VERSION : 0.1
   VAR
      ReadWriteDeviceNo : Int := 0;
      CopyDeviceNO : Int := 0;
      Read : Bool := FALSE;
      Write : Bool := FALSE;
      Copy : Bool := FALSE;
      Tank : Array[0..12] of "UDT502_PV_Tank";
   END_VAR
BEGIN
   Tank[1].Level.PV_Conf_ActV.Address := 324;
   Tank[2].Level.PV_Conf_ActV.Address := 326;
   Tank[1].Level.PV_Conf_ActV.Multiplier := 10.0;
   Tank[2].Level.PV_Conf_ActV.Multiplier := 10.0;
   Tank[1].Level.PV_Conf_ActV.MaxValueSensor := 0.0;
   Tank[2].Level.PV_Conf_ActV.MaxValueSensor := 0.0;
   Tank[2].Level.PV_Conf_ActV.MinValueSensor := 0.0;
   Tank[1].Temp.PV_Conf_ActV.Address := 300;
   Tank[1].Level.PV_Conf_ActV.MinValueSensor := 0.0;
   Tank[2].Temp.PV_Conf_ActV.Address := 302;
   Tank[1].Temp.PV_Conf_ActV.Multiplier := 100.0;
   Tank[2].Temp.PV_Conf_ActV.Multiplier := 100.0;
   Tank[0].Temp.PV_SetV.Value := 15.0;
   Tank[0].Temp.PV_SetV.WarningLowerLimit := 0.0;
   Tank[0].Temp.PV_SetV.WarningUpperLimit := 0.0;
   Tank[0].Temp.PV_SetV.AlarmLowerLimit := 0.0;
   Tank[0].Temp.PV_SetV.AlarmUpperLimit := 0.0;
   Tank[0].Temp.PV_Conf_ActV.ModulNo := 1;
   Tank[0].Temp.PV_Conf_ActV.Address := 300;
   Tank[0].Temp.PV_Conf_ActV.OffsetSignal := 0;
   Tank[0].Temp.PV_Conf_ActV.Multiplier := 100.0;
   Tank[0].Temp.PV_Conf_ActV.MinValueSensor := 1.0;
   Tank[0].Temp.PV_Conf_ActV.MaxValueSensor := 10000.0;
   Tank[0].Temp.PV_Conf_ActV.MaxSignalResolution := 0.0;
   Tank[0].Level.PV_SetV.Value := 0.0;
   Tank[0].Level.PV_SetV.WarningLowerLimit := 0.0;
   Tank[0].Level.PV_SetV.WarningUpperLimit := 0.0;
   Tank[0].Level.PV_SetV.AlarmLowerLimit := 0.0;
   Tank[0].Level.PV_SetV.AlarmUpperLimit := 0.0;
   Tank[0].Level.PV_Conf_ActV.ModulNo := 1;
   Tank[0].Level.PV_Conf_ActV.Address := 324;
   Tank[0].Level.PV_Conf_ActV.OffsetSignal := 0;
   Tank[0].Level.PV_Conf_ActV.Multiplier := 10.0;
   Tank[0].Level.PV_Conf_ActV.MinValueSensor := 0.0;
   Tank[0].Level.PV_Conf_ActV.MaxValueSensor := 0.0;
   Tank[0].Level.PV_Conf_ActV.MaxSignalResolution := 0.0;
   Tank[0].Pressure.PV_SetV.Value := 0.0;
   Tank[0].Pressure.PV_SetV.WarningLowerLimit := 0.0;
   Tank[0].Pressure.PV_SetV.WarningUpperLimit := 0.0;
   Tank[0].Pressure.PV_SetV.AlarmLowerLimit := 0.0;
   Tank[0].Pressure.PV_SetV.AlarmUpperLimit := 0.0;
   Tank[0].Pressure.PV_Conf_ActV.ModulNo := 0;
   Tank[0].Pressure.PV_Conf_ActV.Address := 0;
   Tank[0].Pressure.PV_Conf_ActV.OffsetSignal := 0;
   Tank[0].Pressure.PV_Conf_ActV.Multiplier := 0.0;
   Tank[0].Pressure.PV_Conf_ActV.MinValueSensor := 0.0;
   Tank[0].Pressure.PV_Conf_ActV.MaxValueSensor := 0.0;
   Tank[0].Pressure.PV_Conf_ActV.MaxSignalResolution := 0.0;
   Tank[0].Nucleation.PV_SetV.Value := 2.0;
   Tank[0].Nucleation.PV_SetV.WarningLowerLimit := 0.0;
   Tank[0].Nucleation.PV_SetV.WarningUpperLimit := 0.0;
   Tank[0].Nucleation.PV_SetV.AlarmLowerLimit := 0.0;
   Tank[0].Nucleation.PV_SetV.AlarmUpperLimit := 0.0;
   Tank[0].Nucleation.PV_Conf_ActV.ModulNo := 1;
   Tank[0].Nucleation.PV_Conf_ActV.Address := 330;
   Tank[0].Nucleation.PV_Conf_ActV.OffsetSignal := 0;
   Tank[0].Nucleation.PV_Conf_ActV.Multiplier := 10.0;
   Tank[0].Nucleation.PV_Conf_ActV.MinValueSensor := 0.0;
   Tank[0].Nucleation.PV_Conf_ActV.MaxValueSensor := 100.0;
   Tank[0].Nucleation.PV_Conf_ActV.MaxSignalResolution := 0.0;
   Tank[0].JacketHeater.PV_SetV.Value := 0.0;
   Tank[0].JacketHeater.PV_SetV.WarningLowerLimit := 0.0;
   Tank[0].JacketHeater.PV_SetV.WarningUpperLimit := 0.0;
   Tank[0].JacketHeater.PV_SetV.AlarmLowerLimit := 0.0;
   Tank[0].JacketHeater.PV_SetV.AlarmUpperLimit := 0.0;
   Tank[0].JacketHeater.PV_Conf_ActV.ModulNo := 0;
   Tank[0].JacketHeater.PV_Conf_ActV.Address := 0;
   Tank[0].JacketHeater.PV_Conf_ActV.OffsetSignal := 0;
   Tank[0].JacketHeater.PV_Conf_ActV.Multiplier := 0.0;
   Tank[0].JacketHeater.PV_Conf_ActV.MinValueSensor := 0.0;
   Tank[0].JacketHeater.PV_Conf_ActV.MaxValueSensor := 0.0;
   Tank[0].JacketHeater.PV_Conf_ActV.MaxSignalResolution := 0.0;
   Tank[1].Temp.PV_SetV.Value := 15.0;
   Tank[1].Temp.PV_SetV.WarningLowerLimit := 0.0;
   Tank[1].Temp.PV_SetV.WarningUpperLimit := 0.0;
   Tank[1].Temp.PV_SetV.AlarmLowerLimit := 0.0;
   Tank[1].Temp.PV_SetV.AlarmUpperLimit := 0.0;
   Tank[1].Temp.PV_Conf_ActV.ModulNo := 1;
   Tank[1].Temp.PV_Conf_ActV.OffsetSignal := 0;
   Tank[1].Temp.PV_Conf_ActV.MinValueSensor := 1.0;
   Tank[1].Temp.PV_Conf_ActV.MaxValueSensor := 10000.0;
   Tank[1].Temp.PV_Conf_ActV.MaxSignalResolution := 0.0;
   Tank[1].Level.PV_SetV.Value := 0.0;
   Tank[1].Level.PV_SetV.WarningLowerLimit := 0.0;
   Tank[1].Level.PV_SetV.WarningUpperLimit := 0.0;
   Tank[1].Level.PV_SetV.AlarmLowerLimit := 0.0;
   Tank[1].Level.PV_SetV.AlarmUpperLimit := 0.0;
   Tank[1].Level.PV_Conf_ActV.ModulNo := 1;
   Tank[1].Level.PV_Conf_ActV.OffsetSignal := 0;
   Tank[1].Level.PV_Conf_ActV.MaxSignalResolution := 0.0;
   Tank[1].Pressure.PV_SetV.Value := 0.0;
   Tank[1].Pressure.PV_SetV.WarningLowerLimit := 0.0;
   Tank[1].Pressure.PV_SetV.WarningUpperLimit := 0.0;
   Tank[1].Pressure.PV_SetV.AlarmLowerLimit := 0.0;
   Tank[1].Pressure.PV_SetV.AlarmUpperLimit := 0.0;
   Tank[1].Pressure.PV_Conf_ActV.ModulNo := 0;
   Tank[1].Pressure.PV_Conf_ActV.Address := 0;
   Tank[1].Pressure.PV_Conf_ActV.OffsetSignal := 0;
   Tank[1].Pressure.PV_Conf_ActV.Multiplier := 0.0;
   Tank[1].Pressure.PV_Conf_ActV.MinValueSensor := 0.0;
   Tank[1].Pressure.PV_Conf_ActV.MaxValueSensor := 0.0;
   Tank[1].Pressure.PV_Conf_ActV.MaxSignalResolution := 0.0;
   Tank[1].Nucleation.PV_SetV.Value := 2.0;
   Tank[1].Nucleation.PV_SetV.WarningLowerLimit := 0.0;
   Tank[1].Nucleation.PV_SetV.WarningUpperLimit := 0.0;
   Tank[1].Nucleation.PV_SetV.AlarmLowerLimit := 0.0;
   Tank[1].Nucleation.PV_SetV.AlarmUpperLimit := 0.0;
   Tank[1].Nucleation.PV_Conf_ActV.ModulNo := 1;
   Tank[1].Nucleation.PV_Conf_ActV.Address := 330;
   Tank[1].Nucleation.PV_Conf_ActV.OffsetSignal := 0;
   Tank[1].Nucleation.PV_Conf_ActV.Multiplier := 10.0;
   Tank[1].Nucleation.PV_Conf_ActV.MinValueSensor := 0.0;
   Tank[1].Nucleation.PV_Conf_ActV.MaxValueSensor := 100.0;
   Tank[1].Nucleation.PV_Conf_ActV.MaxSignalResolution := 0.0;
   Tank[1].JacketHeater.PV_SetV.Value := 0.0;
   Tank[1].JacketHeater.PV_SetV.WarningLowerLimit := 0.0;
   Tank[1].JacketHeater.PV_SetV.WarningUpperLimit := 0.0;
   Tank[1].JacketHeater.PV_SetV.AlarmLowerLimit := 0.0;
   Tank[1].JacketHeater.PV_SetV.AlarmUpperLimit := 0.0;
   Tank[1].JacketHeater.PV_Conf_ActV.ModulNo := 0;
   Tank[1].JacketHeater.PV_Conf_ActV.Address := 0;
   Tank[1].JacketHeater.PV_Conf_ActV.OffsetSignal := 0;
   Tank[1].JacketHeater.PV_Conf_ActV.Multiplier := 0.0;
   Tank[1].JacketHeater.PV_Conf_ActV.MinValueSensor := 0.0;
   Tank[1].JacketHeater.PV_Conf_ActV.MaxValueSensor := 0.0;
   Tank[1].JacketHeater.PV_Conf_ActV.MaxSignalResolution := 0.0;
   Tank[2].Temp.PV_SetV.Value := 15.0;
   Tank[2].Temp.PV_SetV.WarningLowerLimit := 0.0;
   Tank[2].Temp.PV_SetV.WarningUpperLimit := 0.0;
   Tank[2].Temp.PV_SetV.AlarmLowerLimit := 0.0;
   Tank[2].Temp.PV_SetV.AlarmUpperLimit := 0.0;
   Tank[2].Temp.PV_Conf_ActV.ModulNo := 1;
   Tank[2].Temp.PV_Conf_ActV.OffsetSignal := 0;
   Tank[2].Temp.PV_Conf_ActV.MinValueSensor := 1.0;
   Tank[2].Temp.PV_Conf_ActV.MaxValueSensor := 10000.0;
   Tank[2].Temp.PV_Conf_ActV.MaxSignalResolution := 0.0;
   Tank[2].Level.PV_SetV.Value := 0.0;
   Tank[2].Level.PV_SetV.WarningLowerLimit := 0.0;
   Tank[2].Level.PV_SetV.WarningUpperLimit := 0.0;
   Tank[2].Level.PV_SetV.AlarmLowerLimit := 0.0;
   Tank[2].Level.PV_SetV.AlarmUpperLimit := 0.0;
   Tank[2].Level.PV_Conf_ActV.ModulNo := 1;
   Tank[2].Level.PV_Conf_ActV.OffsetSignal := 0;
   Tank[2].Level.PV_Conf_ActV.MaxSignalResolution := 0.0;
   Tank[2].Pressure.PV_SetV.Value := 0.0;
   Tank[2].Pressure.PV_SetV.WarningLowerLimit := 0.0;
   Tank[2].Pressure.PV_SetV.WarningUpperLimit := 0.0;
   Tank[2].Pressure.PV_SetV.AlarmLowerLimit := 0.0;
   Tank[2].Pressure.PV_SetV.AlarmUpperLimit := 0.0;
   Tank[2].Pressure.PV_Conf_ActV.ModulNo := 0;
   Tank[2].Pressure.PV_Conf_ActV.Address := 0;
   Tank[2].Pressure.PV_Conf_ActV.OffsetSignal := 0;
   Tank[2].Pressure.PV_Conf_ActV.Multiplier := 0.0;
   Tank[2].Pressure.PV_Conf_ActV.MinValueSensor := 0.0;
   Tank[2].Pressure.PV_Conf_ActV.MaxValueSensor := 0.0;
   Tank[2].Pressure.PV_Conf_ActV.MaxSignalResolution := 0.0;
   Tank[2].Nucleation.PV_SetV.Value := 0.0;
   Tank[2].Nucleation.PV_SetV.WarningLowerLimit := 0.0;
   Tank[2].Nucleation.PV_SetV.WarningUpperLimit := 0.0;
   Tank[2].Nucleation.PV_SetV.AlarmLowerLimit := 0.0;
   Tank[2].Nucleation.PV_SetV.AlarmUpperLimit := 0.0;
   Tank[2].Nucleation.PV_Conf_ActV.ModulNo := 0;
   Tank[2].Nucleation.PV_Conf_ActV.Address := 0;
   Tank[2].Nucleation.PV_Conf_ActV.OffsetSignal := 0;
   Tank[2].Nucleation.PV_Conf_ActV.Multiplier := 10.0;
   Tank[2].Nucleation.PV_Conf_ActV.MinValueSensor := 0.0;
   Tank[2].Nucleation.PV_Conf_ActV.MaxValueSensor := 0.0;
   Tank[2].Nucleation.PV_Conf_ActV.MaxSignalResolution := 0.0;
   Tank[2].JacketHeater.PV_SetV.Value := 0.0;
   Tank[2].JacketHeater.PV_SetV.WarningLowerLimit := 0.0;
   Tank[2].JacketHeater.PV_SetV.WarningUpperLimit := 0.0;
   Tank[2].JacketHeater.PV_SetV.AlarmLowerLimit := 0.0;
   Tank[2].JacketHeater.PV_SetV.AlarmUpperLimit := 0.0;
   Tank[2].JacketHeater.PV_Conf_ActV.ModulNo := 0;
   Tank[2].JacketHeater.PV_Conf_ActV.Address := 0;
   Tank[2].JacketHeater.PV_Conf_ActV.OffsetSignal := 0;
   Tank[2].JacketHeater.PV_Conf_ActV.Multiplier := 0.0;
   Tank[2].JacketHeater.PV_Conf_ActV.MinValueSensor := 0.0;
   Tank[2].JacketHeater.PV_Conf_ActV.MaxValueSensor := 0.0;
   Tank[2].JacketHeater.PV_Conf_ActV.MaxSignalResolution := 0.0;
   Tank[3].Temp.PV_SetV.Value := 0.0;
   Tank[3].Temp.PV_SetV.WarningLowerLimit := 0.0;
   Tank[3].Temp.PV_SetV.WarningUpperLimit := 0.0;
   Tank[3].Temp.PV_SetV.AlarmLowerLimit := 0.0;
   Tank[3].Temp.PV_SetV.AlarmUpperLimit := 0.0;
   Tank[3].Temp.PV_Conf_ActV.ModulNo := 0;
   Tank[3].Temp.PV_Conf_ActV.Address := 516;
   Tank[3].Temp.PV_Conf_ActV.OffsetSignal := 0;
   Tank[3].Temp.PV_Conf_ActV.Multiplier := 10.0;
   Tank[3].Temp.PV_Conf_ActV.MinValueSensor := 0.0;
   Tank[3].Temp.PV_Conf_ActV.MaxValueSensor := 0.0;
   Tank[3].Temp.PV_Conf_ActV.MaxSignalResolution := 0.0;
   Tank[3].Level.PV_SetV.Value := 0.0;
   Tank[3].Level.PV_SetV.WarningLowerLimit := 0.0;
   Tank[3].Level.PV_SetV.WarningUpperLimit := 0.0;
   Tank[3].Level.PV_SetV.AlarmLowerLimit := 0.0;
   Tank[3].Level.PV_SetV.AlarmUpperLimit := 0.0;
   Tank[3].Level.PV_Conf_ActV.ModulNo := 0;
   Tank[3].Level.PV_Conf_ActV.Address := 0;
   Tank[3].Level.PV_Conf_ActV.OffsetSignal := 0;
   // 710 more start values not shown
END_DATA_BLOCK

DATA_BLOCK "DB604_PV_Mixinghead"   // DB604
TITLE = Process values of mixinghead
{ S7_Optimized_Access := 'FALSE' }
AUTHOR : KT242
VERSION : 0.1
   VAR
      ReadWriteDeviceNo : Int := 0;
      CopyDeviceNO : Int := 0;
      Read : Bool := FALSE;
      Write : Bool := FALSE;
      Copy : Bool := FALSE;
      Mixinghead : Array[0..16] of "UDT504_PV_MH";   // Process value of the mixinghead 1 - 16
   END_VAR
BEGIN
   Mixinghead[0].Pressure_Connection[1].PV_SetV.Value := 120.0;
   Mixinghead[0].Pressure_Connection[1].PV_SetV.WarningLowerLimit := 0.0;
   Mixinghead[0].Pressure_Connection[1].PV_SetV.WarningUpperLimit := 0.0;
   Mixinghead[0].Pressure_Connection[1].PV_SetV.AlarmLowerLimit := 0.0;
   Mixinghead[0].Pressure_Connection[1].PV_SetV.AlarmUpperLimit := 0.0;
   Mixinghead[0].Pressure_Connection[1].PV_ActV.Value := 3.2;
   Mixinghead[0].Pressure_Connection[1].PV_ActV.ValueState := 16#0000;
   Mixinghead[0].Pressure_Connection[1].PV_Conf_ActV.ModulNo := 2;
   Mixinghead[0].Pressure_Connection[1].PV_Conf_ActV.Address := 412;
   Mixinghead[0].Pressure_Connection[1].PV_Conf_ActV.OffsetSignal := 0;
   Mixinghead[0].Pressure_Connection[1].PV_Conf_ActV.Multiplier := 10.0;
   Mixinghead[0].Pressure_Connection[1].PV_Conf_ActV.MinValueSensor := -50.0;
   Mixinghead[0].Pressure_Connection[1].PV_Conf_ActV.MaxValueSensor := 60000.0;
   Mixinghead[0].Pressure_Connection[1].PV_Conf_ActV.MaxSignalResolution := 0.0;
   Mixinghead[0].Pressure_Connection[2].PV_SetV.Value := 120.0;
   Mixinghead[0].Pressure_Connection[2].PV_SetV.WarningLowerLimit := 0.0;
   Mixinghead[0].Pressure_Connection[2].PV_SetV.WarningUpperLimit := 0.0;
   Mixinghead[0].Pressure_Connection[2].PV_SetV.AlarmLowerLimit := 0.0;
   Mixinghead[0].Pressure_Connection[2].PV_SetV.AlarmUpperLimit := 0.0;
   Mixinghead[0].Pressure_Connection[2].PV_ActV.Value := 2.4;
   Mixinghead[0].Pressure_Connection[2].PV_ActV.ValueState := 16#0000;
   Mixinghead[0].Pressure_Connection[2].PV_Conf_ActV.ModulNo := 2;
   Mixinghead[0].Pressure_Connection[2].PV_Conf_ActV.Address := 414;
   Mixinghead[0].Pressure_Connection[2].PV_Conf_ActV.OffsetSignal := 0;
   Mixinghead[0].Pressure_Connection[2].PV_Conf_ActV.Multiplier := 10.0;
   Mixinghead[0].Pressure_Connection[2].PV_Conf_ActV.MinValueSensor := -50.0;
   Mixinghead[0].Pressure_Connection[2].PV_Conf_ActV.MaxValueSensor := 60000.0;
   Mixinghead[0].Pressure_Connection[2].PV_Conf_ActV.MaxSignalResolution := 0.0;
   Mixinghead[0].Pressure_Connection[3].PV_SetV.Value := 0.0;
   Mixinghead[0].Pressure_Connection[3].PV_SetV.WarningLowerLimit := 0.0;
   Mixinghead[0].Pressure_Connection[3].PV_SetV.WarningUpperLimit := 0.0;
   Mixinghead[0].Pressure_Connection[3].PV_SetV.AlarmLowerLimit := 0.0;
   Mixinghead[0].Pressure_Connection[3].PV_SetV.AlarmUpperLimit := 0.0;
   Mixinghead[0].Pressure_Connection[3].PV_ActV.Value := 0.0;
   Mixinghead[0].Pressure_Connection[3].PV_ActV.ValueState := 16#0000;
   Mixinghead[0].Pressure_Connection[3].PV_Conf_ActV.ModulNo := 0;
   Mixinghead[0].Pressure_Connection[3].PV_Conf_ActV.Address := 0;
   Mixinghead[0].Pressure_Connection[3].PV_Conf_ActV.OffsetSignal := 0;
   Mixinghead[0].Pressure_Connection[3].PV_Conf_ActV.Multiplier := 0.0;
   Mixinghead[0].Pressure_Connection[3].PV_Conf_ActV.MinValueSensor := 0.0;
   Mixinghead[0].Pressure_Connection[3].PV_Conf_ActV.MaxValueSensor := 0.0;
   Mixinghead[0].Pressure_Connection[3].PV_Conf_ActV.MaxSignalResolution := 0.0;
   Mixinghead[0].Pressure_Connection[4].PV_SetV.Value := 0.0;
   Mixinghead[0].Pressure_Connection[4].PV_SetV.WarningLowerLimit := 0.0;
   Mixinghead[0].Pressure_Connection[4].PV_SetV.WarningUpperLimit := 0.0;
   Mixinghead[0].Pressure_Connection[4].PV_SetV.AlarmLowerLimit := 0.0;
   Mixinghead[0].Pressure_Connection[4].PV_SetV.AlarmUpperLimit := 0.0;
   Mixinghead[0].Pressure_Connection[4].PV_ActV.Value := 0.0;
   Mixinghead[0].Pressure_Connection[4].PV_ActV.ValueState := 16#0000;
   Mixinghead[0].Pressure_Connection[4].PV_Conf_ActV.ModulNo := 0;
   Mixinghead[0].Pressure_Connection[4].PV_Conf_ActV.Address := 0;
   Mixinghead[0].Pressure_Connection[4].PV_Conf_ActV.OffsetSignal := 0;
   Mixinghead[0].Pressure_Connection[4].PV_Conf_ActV.Multiplier := 0.0;
   Mixinghead[0].Pressure_Connection[4].PV_Conf_ActV.MinValueSensor := 0.0;
   Mixinghead[0].Pressure_Connection[4].PV_Conf_ActV.MaxValueSensor := 0.0;
   Mixinghead[0].Pressure_Connection[4].PV_Conf_ActV.MaxSignalResolution := 0.0;
   Mixinghead[0].Pressure_Connection[5].PV_SetV.Value := 0.0;
   Mixinghead[0].Pressure_Connection[5].PV_SetV.WarningLowerLimit := 0.0;
   Mixinghead[0].Pressure_Connection[5].PV_SetV.WarningUpperLimit := 0.0;
   Mixinghead[0].Pressure_Connection[5].PV_SetV.AlarmLowerLimit := 0.0;
   Mixinghead[0].Pressure_Connection[5].PV_SetV.AlarmUpperLimit := 0.0;
   Mixinghead[0].Pressure_Connection[5].PV_ActV.Value := 0.0;
   Mixinghead[0].Pressure_Connection[5].PV_ActV.ValueState := 16#0000;
   Mixinghead[0].Pressure_Connection[5].PV_Conf_ActV.ModulNo := 0;
   Mixinghead[0].Pressure_Connection[5].PV_Conf_ActV.Address := 0;
   Mixinghead[0].Pressure_Connection[5].PV_Conf_ActV.OffsetSignal := 0;
   Mixinghead[0].Pressure_Connection[5].PV_Conf_ActV.Multiplier := 0.0;
   Mixinghead[0].Pressure_Connection[5].PV_Conf_ActV.MinValueSensor := 0.0;
   Mixinghead[0].Pressure_Connection[5].PV_Conf_ActV.MaxValueSensor := 0.0;
   Mixinghead[0].Pressure_Connection[5].PV_Conf_ActV.MaxSignalResolution := 0.0;
   Mixinghead[0].Pressure_Connection[6].PV_SetV.Value := 0.0;
   Mixinghead[0].Pressure_Connection[6].PV_SetV.WarningLowerLimit := 0.0;
   Mixinghead[0].Pressure_Connection[6].PV_SetV.WarningUpperLimit := 0.0;
   Mixinghead[0].Pressure_Connection[6].PV_SetV.AlarmLowerLimit := 0.0;
   Mixinghead[0].Pressure_Connection[6].PV_SetV.AlarmUpperLimit := 0.0;
   Mixinghead[0].Pressure_Connection[6].PV_ActV.Value := 0.0;
   Mixinghead[0].Pressure_Connection[6].PV_ActV.ValueState := 16#0000;
   Mixinghead[0].Pressure_Connection[6].PV_Conf_ActV.ModulNo := 0;
   Mixinghead[0].Pressure_Connection[6].PV_Conf_ActV.Address := 0;
   Mixinghead[0].Pressure_Connection[6].PV_Conf_ActV.OffsetSignal := 0;
   Mixinghead[0].Pressure_Connection[6].PV_Conf_ActV.Multiplier := 0.0;
   Mixinghead[0].Pressure_Connection[6].PV_Conf_ActV.MinValueSensor := 0.0;
   Mixinghead[0].Pressure_Connection[6].PV_Conf_ActV.MaxValueSensor := 0.0;
   Mixinghead[0].Pressure_Connection[6].PV_Conf_ActV.MaxSignalResolution := 0.0;
   Mixinghead[0].Temperature_Connection[1].PV_SetV.Value := 0.0;
   Mixinghead[0].Temperature_Connection[1].PV_SetV.WarningLowerLimit := 0.0;
   Mixinghead[0].Temperature_Connection[1].PV_SetV.WarningUpperLimit := 0.0;
   Mixinghead[0].Temperature_Connection[1].PV_SetV.AlarmLowerLimit := 0.0;
   Mixinghead[0].Temperature_Connection[1].PV_SetV.AlarmUpperLimit := 0.0;
   Mixinghead[0].Temperature_Connection[1].PV_ActV.Value := 26.26;
   Mixinghead[0].Temperature_Connection[1].PV_ActV.ValueState := 16#0000;
   Mixinghead[0].Temperature_Connection[1].PV_Conf_ActV.ModulNo := 2;
   Mixinghead[0].Temperature_Connection[1].PV_Conf_ActV.Address := 396;
   Mixinghead[0].Temperature_Connection[1].PV_Conf_ActV.OffsetSignal := 0;
   Mixinghead[0].Temperature_Connection[1].PV_Conf_ActV.Multiplier := 100.0;
   Mixinghead[0].Temperature_Connection[1].PV_Conf_ActV.MinValueSensor := 1.0;
   Mixinghead[0].Temperature_Connection[1].PV_Conf_ActV.MaxValueSensor := 10000.0;
   Mixinghead[0].Temperature_Connection[1].PV_Conf_ActV.MaxSignalResolution := 0.0;
   Mixinghead[0].Temperature_Connection[2].PV_SetV.Value := 0.0;
   Mixinghead[0].Temperature_Connection[2].PV_SetV.WarningLowerLimit := 0.0;
   Mixinghead[0].Temperature_Connection[2].PV_SetV.WarningUpperLimit := 0.0;
   Mixinghead[0].Temperature_Connection[2].PV_SetV.AlarmLowerLimit := 0.0;
   Mixinghead[0].Temperature_Connection[2].PV_SetV.AlarmUpperLimit := 0.0;
   Mixinghead[0].Temperature_Connection[2].PV_ActV.Value := 25.85;
   Mixinghead[0].Temperature_Connection[2].PV_ActV.ValueState := 16#0000;
   Mixinghead[0].Temperature_Connection[2].PV_Conf_ActV.ModulNo := 2;
   Mixinghead[0].Temperature_Connection[2].PV_Conf_ActV.Address := 398;
   Mixinghead[0].Temperature_Connection[2].PV_Conf_ActV.OffsetSignal := 0;
   Mixinghead[0].Temperature_Connection[2].PV_Conf_ActV.Multiplier := 100.0;
   Mixinghead[0].Temperature_Connection[2].PV_Conf_ActV.MinValueSensor := 1.0;
   Mixinghead[0].Temperature_Connection[2].PV_Conf_ActV.MaxValueSensor := 10000.0;
   Mixinghead[0].Temperature_Connection[2].PV_Conf_ActV.MaxSignalResolution := 0.0;
   Mixinghead[0].Temperature_Connection[3].PV_SetV.Value := 0.0;
   Mixinghead[0].Temperature_Connection[3].PV_SetV.WarningLowerLimit := 0.0;
   Mixinghead[0].Temperature_Connection[3].PV_SetV.WarningUpperLimit := 0.0;
   Mixinghead[0].Temperature_Connection[3].PV_SetV.AlarmLowerLimit := 0.0;
   Mixinghead[0].Temperature_Connection[3].PV_SetV.AlarmUpperLimit := 0.0;
   Mixinghead[0].Temperature_Connection[3].PV_ActV.Value := 0.0;
   Mixinghead[0].Temperature_Connection[3].PV_ActV.ValueState := 16#0000;
   Mixinghead[0].Temperature_Connection[3].PV_Conf_ActV.ModulNo := 0;
   Mixinghead[0].Temperature_Connection[3].PV_Conf_ActV.Address := 0;
   Mixinghead[0].Temperature_Connection[3].PV_Conf_ActV.OffsetSignal := 0;
   Mixinghead[0].Temperature_Connection[3].PV_Conf_ActV.Multiplier := 0.0;
   Mixinghead[0].Temperature_Connection[3].PV_Conf_ActV.MinValueSensor := 0.0;
   Mixinghead[0].Temperature_Connection[3].PV_Conf_ActV.MaxValueSensor := 0.0;
   Mixinghead[0].Temperature_Connection[3].PV_Conf_ActV.MaxSignalResolution := 0.0;
   Mixinghead[0].Temperature_Connection[4].PV_SetV.Value := 0.0;
   Mixinghead[0].Temperature_Connection[4].PV_SetV.WarningLowerLimit := 0.0;
   Mixinghead[0].Temperature_Connection[4].PV_SetV.WarningUpperLimit := 0.0;
   Mixinghead[0].Temperature_Connection[4].PV_SetV.AlarmLowerLimit := 0.0;
   Mixinghead[0].Temperature_Connection[4].PV_SetV.AlarmUpperLimit := 0.0;
   Mixinghead[0].Temperature_Connection[4].PV_ActV.Value := 0.0;
   Mixinghead[0].Temperature_Connection[4].PV_ActV.ValueState := 16#0000;
   Mixinghead[0].Temperature_Connection[4].PV_Conf_ActV.ModulNo := 0;
   Mixinghead[0].Temperature_Connection[4].PV_Conf_ActV.Address := 0;
   Mixinghead[0].Temperature_Connection[4].PV_Conf_ActV.OffsetSignal := 0;
   Mixinghead[0].Temperature_Connection[4].PV_Conf_ActV.Multiplier := 0.0;
   Mixinghead[0].Temperature_Connection[4].PV_Conf_ActV.MinValueSensor := 0.0;
   Mixinghead[0].Temperature_Connection[4].PV_Conf_ActV.MaxValueSensor := 0.0;
   Mixinghead[0].Temperature_Connection[4].PV_Conf_ActV.MaxSignalResolution := 0.0;
   Mixinghead[0].Temperature_Connection[5].PV_SetV.Value := 0.0;
   Mixinghead[0].Temperature_Connection[5].PV_SetV.WarningLowerLimit := 0.0;
   Mixinghead[0].Temperature_Connection[5].PV_SetV.WarningUpperLimit := 0.0;
   Mixinghead[0].Temperature_Connection[5].PV_SetV.AlarmLowerLimit := 0.0;
   Mixinghead[0].Temperature_Connection[5].PV_SetV.AlarmUpperLimit := 0.0;
   Mixinghead[0].Temperature_Connection[5].PV_ActV.Value := 0.0;
   Mixinghead[0].Temperature_Connection[5].PV_ActV.ValueState := 16#0000;
   Mixinghead[0].Temperature_Connection[5].PV_Conf_ActV.ModulNo := 0;
   Mixinghead[0].Temperature_Connection[5].PV_Conf_ActV.Address := 0;
   Mixinghead[0].Temperature_Connection[5].PV_Conf_ActV.OffsetSignal := 0;
   Mixinghead[0].Temperature_Connection[5].PV_Conf_ActV.Multiplier := 0.0;
   Mixinghead[0].Temperature_Connection[5].PV_Conf_ActV.MinValueSensor := 0.0;
   Mixinghead[0].Temperature_Connection[5].PV_Conf_ActV.MaxValueSensor := 0.0;
   Mixinghead[0].Temperature_Connection[5].PV_Conf_ActV.MaxSignalResolution := 0.0;
   Mixinghead[0].Temperature_Connection[6].PV_SetV.Value := 0.0;
   Mixinghead[0].Temperature_Connection[6].PV_SetV.WarningLowerLimit := 0.0;
   Mixinghead[0].Temperature_Connection[6].PV_SetV.WarningUpperLimit := 0.0;
   Mixinghead[0].Temperature_Connection[6].PV_SetV.AlarmLowerLimit := 0.0;
   Mixinghead[0].Temperature_Connection[6].PV_SetV.AlarmUpperLimit := 0.0;
   Mixinghead[0].Temperature_Connection[6].PV_ActV.Value := 0.0;
   Mixinghead[0].Temperature_Connection[6].PV_ActV.ValueState := 16#0000;
   Mixinghead[0].Temperature_Connection[6].PV_Conf_ActV.ModulNo := 0;
   Mixinghead[0].Temperature_Connection[6].PV_Conf_ActV.Address := 0;
   Mixinghead[0].Temperature_Connection[6].PV_Conf_ActV.OffsetSignal := 0;
   Mixinghead[0].Temperature_Connection[6].PV_Conf_ActV.Multiplier := 0.0;
   Mixinghead[0].Temperature_Connection[6].PV_Conf_ActV.MinValueSensor := 0.0;
   Mixinghead[0].Temperature_Connection[6].PV_Conf_ActV.MaxValueSensor := 0.0;
   Mixinghead[0].Temperature_Connection[6].PV_Conf_ActV.MaxSignalResolution := 0.0;
   Mixinghead[0].SteeringPiston.PV_SetV.Value := 0.0;
   Mixinghead[0].SteeringPiston.PV_SetV.WarningLowerLimit := 0.0;
   Mixinghead[0].SteeringPiston.PV_SetV.WarningUpperLimit := 0.0;
   Mixinghead[0].SteeringPiston.PV_SetV.AlarmLowerLimit := 0.0;
   Mixinghead[0].SteeringPiston.PV_SetV.AlarmUpperLimit := 0.0;
   Mixinghead[0].SteeringPiston.PV_ActV.Value := 0.0;
   Mixinghead[0].SteeringPiston.PV_ActV.ValueState := 16#0000;
   Mixinghead[0].SteeringPiston.PV_Conf_ActV.ModulNo := 0;
   Mixinghead[0].SteeringPiston.PV_Conf_ActV.Address := 0;
   Mixinghead[0].SteeringPiston.PV_Conf_ActV.OffsetSignal := 0;
   Mixinghead[0].SteeringPiston.PV_Conf_ActV.Multiplier := 0.0;
   Mixinghead[0].SteeringPiston.PV_Conf_ActV.MinValueSensor := 0.0;
   Mixinghead[0].SteeringPiston.PV_Conf_ActV.MaxValueSensor := 0.0;
   Mixinghead[0].SteeringPiston.PV_Conf_ActV.MaxSignalResolution := 0.0;
   Mixinghead[0].Inerting.PV_SetV.Value := 0.0;
   Mixinghead[0].Inerting.PV_SetV.WarningLowerLimit := 0.0;
   Mixinghead[0].Inerting.PV_SetV.WarningUpperLimit := 0.0;
   Mixinghead[0].Inerting.PV_SetV.AlarmLowerLimit := 0.0;
   Mixinghead[0].Inerting.PV_SetV.AlarmUpperLimit := 0.0;
   Mixinghead[0].Inerting.PV_ActV.Value := 0.0;
   Mixinghead[0].Inerting.PV_ActV.ValueState := 16#0000;
   Mixinghead[0].Inerting.PV_Conf_ActV.ModulNo := 2;
   Mixinghead[0].Inerting.PV_Conf_ActV.Address := 0;
   Mixinghead[0].Inerting.PV_Conf_ActV.OffsetSignal := 0;
   Mixinghead[0].Inerting.PV_Conf_ActV.Multiplier := 10.0;
   Mixinghead[0].Inerting.PV_Conf_ActV.MinValueSensor := 0.0;
   Mixinghead[0].Inerting.PV_Conf_ActV.MaxValueSensor := 0.0;
   Mixinghead[0].Inerting.PV_Conf_ActV.MaxSignalResolution := 0.0;
   Mixinghead[1].Pressure_Connection[1].PV_SetV.Value := 120.0;
   Mixinghead[1].Pressure_Connection[1].PV_SetV.WarningLowerLimit := 0.0;
   Mixinghead[1].Pressure_Connection[1].PV_SetV.WarningUpperLimit := 0.0;
   Mixinghead[1].Pressure_Connection[1].PV_SetV.AlarmLowerLimit := 0.0;
   // 3370 more start values not shown
END_DATA_BLOCK

DATA_BLOCK "DB606_PV_Machine"   // DB606
TITLE = Process values of machine
{ S7_Optimized_Access := 'FALSE' }
AUTHOR : KT242
VERSION : 0.1
   VAR
      Machine : Array[0..2] of "UDT506_PV_Machine";
   END_VAR
BEGIN
   Machine[0].ShotTime.PV_SetV.Value := 0.0;
   Machine[0].ShotTime.PV_SetV.WarningLowerLimit := 0.0;
   Machine[0].ShotTime.PV_SetV.WarningUpperLimit := 0.0;
   Machine[0].ShotTime.PV_SetV.AlarmLowerLimit := 0.0;
   Machine[0].ShotTime.PV_SetV.AlarmUpperLimit := 0.0;
   Machine[0].ShotTime.PV_ActV.Value := 0.0;
   Machine[0].ShotTime.PV_ActV.ValueState := 16#0000;
   Machine[0].ShotTime.PV_Conf_ActV.ModulNo := 0;
   Machine[0].ShotTime.PV_Conf_ActV.Address := 0;
   Machine[0].ShotTime.PV_Conf_ActV.OffsetSignal := 0;
   Machine[0].ShotTime.PV_Conf_ActV.Multiplier := 0.0;
   Machine[0].ShotTime.PV_Conf_ActV.MinValueSensor := 0.0;
   Machine[0].ShotTime.PV_Conf_ActV.MaxValueSensor := 0.0;
   Machine[0].ShotTime.PV_Conf_ActV.MaxSignalResolution := 0.0;
   Machine[0].Discharge.PV_SetV.Value := 0.0;
   Machine[0].Discharge.PV_SetV.WarningLowerLimit := 0.0;
   Machine[0].Discharge.PV_SetV.WarningUpperLimit := 0.0;
   Machine[0].Discharge.PV_SetV.AlarmLowerLimit := 0.0;
   Machine[0].Discharge.PV_SetV.AlarmUpperLimit := 0.0;
   Machine[0].Discharge.PV_ActV.Value := 0.0;
   Machine[0].Discharge.PV_ActV.ValueState := 16#0000;
   Machine[0].Discharge.PV_Conf_ActV.ModulNo := 0;
   Machine[0].Discharge.PV_Conf_ActV.Address := 0;
   Machine[0].Discharge.PV_Conf_ActV.OffsetSignal := 0;
   Machine[0].Discharge.PV_Conf_ActV.Multiplier := 0.0;
   Machine[0].Discharge.PV_Conf_ActV.MinValueSensor := 0.0;
   Machine[0].Discharge.PV_Conf_ActV.MaxValueSensor := 0.0;
   Machine[0].Discharge.PV_Conf_ActV.MaxSignalResolution := 0.0;
   Machine[1].ShotTime.PV_SetV.Value := 100.0;
   Machine[1].ShotTime.PV_SetV.WarningLowerLimit := 0.0;
   Machine[1].ShotTime.PV_SetV.WarningUpperLimit := 0.0;
   Machine[1].ShotTime.PV_SetV.AlarmLowerLimit := 0.0;
   Machine[1].ShotTime.PV_SetV.AlarmUpperLimit := 0.0;
   Machine[1].ShotTime.PV_ActV.Value := 0.964;
   Machine[1].ShotTime.PV_ActV.ValueState := 16#0000;
   Machine[1].ShotTime.PV_Conf_ActV.ModulNo := 0;
   Machine[1].ShotTime.PV_Conf_ActV.Address := 0;
   Machine[1].ShotTime.PV_Conf_ActV.OffsetSignal := 0;
   Machine[1].ShotTime.PV_Conf_ActV.Multiplier := 0.0;
   Machine[1].ShotTime.PV_Conf_ActV.MinValueSensor := 0.0;
   Machine[1].ShotTime.PV_Conf_ActV.MaxValueSensor := 0.0;
   Machine[1].ShotTime.PV_Conf_ActV.MaxSignalResolution := 0.0;
   Machine[1].Discharge.PV_SetV.Value := 0.0;
   Machine[1].Discharge.PV_SetV.WarningLowerLimit := 0.0;
   Machine[1].Discharge.PV_SetV.WarningUpperLimit := 0.0;
   Machine[1].Discharge.PV_SetV.AlarmLowerLimit := 0.0;
   Machine[1].Discharge.PV_SetV.AlarmUpperLimit := 0.0;
   Machine[1].Discharge.PV_ActV.Value := 0.0;
   Machine[1].Discharge.PV_ActV.ValueState := 16#0000;
   Machine[1].Discharge.PV_Conf_ActV.ModulNo := 0;
   Machine[1].Discharge.PV_Conf_ActV.Address := 0;
   Machine[1].Discharge.PV_Conf_ActV.OffsetSignal := 0;
   Machine[1].Discharge.PV_Conf_ActV.Multiplier := 0.0;
   Machine[1].Discharge.PV_Conf_ActV.MinValueSensor := 0.0;
   Machine[1].Discharge.PV_Conf_ActV.MaxValueSensor := 0.0;
   Machine[1].Discharge.PV_Conf_ActV.MaxSignalResolution := 0.0;
   Machine[2].ShotTime.PV_SetV.Value := 0.0;
   Machine[2].ShotTime.PV_SetV.WarningLowerLimit := 0.0;
   Machine[2].ShotTime.PV_SetV.WarningUpperLimit := 0.0;
   Machine[2].ShotTime.PV_SetV.AlarmLowerLimit := 0.0;
   Machine[2].ShotTime.PV_SetV.AlarmUpperLimit := 0.0;
   Machine[2].ShotTime.PV_ActV.Value := 0.0;
   Machine[2].ShotTime.PV_ActV.ValueState := 16#0000;
   Machine[2].ShotTime.PV_Conf_ActV.ModulNo := 0;
   Machine[2].ShotTime.PV_Conf_ActV.Address := 0;
   Machine[2].ShotTime.PV_Conf_ActV.OffsetSignal := 0;
   Machine[2].ShotTime.PV_Conf_ActV.Multiplier := 0.0;
   Machine[2].ShotTime.PV_Conf_ActV.MinValueSensor := 0.0;
   Machine[2].ShotTime.PV_Conf_ActV.MaxValueSensor := 0.0;
   Machine[2].ShotTime.PV_Conf_ActV.MaxSignalResolution := 0.0;
   Machine[2].Discharge.PV_SetV.Value := 0.0;
   Machine[2].Discharge.PV_SetV.WarningLowerLimit := 0.0;
   Machine[2].Discharge.PV_SetV.WarningUpperLimit := 0.0;
   Machine[2].Discharge.PV_SetV.AlarmLowerLimit := 0.0;
   Machine[2].Discharge.PV_SetV.AlarmUpperLimit := 0.0;
   Machine[2].Discharge.PV_ActV.Value := 0.0;
   Machine[2].Discharge.PV_ActV.ValueState := 16#0000;
   Machine[2].Discharge.PV_Conf_ActV.ModulNo := 0;
   Machine[2].Discharge.PV_Conf_ActV.Address := 0;
   Machine[2].Discharge.PV_Conf_ActV.OffsetSignal := 0;
   Machine[2].Discharge.PV_Conf_ActV.Multiplier := 0.0;
   Machine[2].Discharge.PV_Conf_ActV.MinValueSensor := 0.0;
   Machine[2].Discharge.PV_Conf_ActV.MaxValueSensor := 0.0;
   Machine[2].Discharge.PV_Conf_ActV.MaxSignalResolution := 0.0;
   Machine[1].PneumaticFlow.PV_Conf_ActV.ModulNo := 1;
   Machine[1].PneumaticFlow.PV_Conf_ActV.Address := 330;
   Machine[1].PneumaticFlow.PV_Conf_ActV.Multiplier := 1.18;
   Machine[1].PneumaticFlow.PV_Conf_ActV.MinValueSensor := 5.0;
   Machine[1].PneumaticFlow.PV_Conf_ActV.MaxValueSensor := 5000.0;
   Machine[0].PneumaticFlow.PV_SetV.Value := 0.0;
   Machine[0].PneumaticFlow.PV_SetV.WarningLowerLimit := 0.0;
   Machine[0].PneumaticFlow.PV_SetV.WarningUpperLimit := 0.0;
   Machine[0].PneumaticFlow.PV_SetV.AlarmLowerLimit := 0.0;
   Machine[0].PneumaticFlow.PV_SetV.AlarmUpperLimit := 0.0;
   Machine[0].PneumaticFlow.PV_ActV.Value := 0.0;
   Machine[0].PneumaticFlow.PV_ActV.ValueState := 16#0000;
   Machine[0].PneumaticFlow.PV_Conf_ActV.ModulNo := 0;
   Machine[0].PneumaticFlow.PV_Conf_ActV.Address := 0;
   Machine[0].PneumaticFlow.PV_Conf_ActV.OffsetSignal := 0;
   Machine[0].PneumaticFlow.PV_Conf_ActV.Multiplier := 0.0;
   Machine[0].PneumaticFlow.PV_Conf_ActV.MinValueSensor := 0.0;
   Machine[0].PneumaticFlow.PV_Conf_ActV.MaxValueSensor := 0.0;
   Machine[0].PneumaticFlow.PV_Conf_ActV.MaxSignalResolution := 0.0;
   Machine[1].PneumaticFlow.PV_SetV.Value := 0.0;
   Machine[1].PneumaticFlow.PV_SetV.WarningLowerLimit := 0.0;
   Machine[1].PneumaticFlow.PV_SetV.WarningUpperLimit := 0.0;
   Machine[1].PneumaticFlow.PV_SetV.AlarmLowerLimit := 0.0;
   Machine[1].PneumaticFlow.PV_SetV.AlarmUpperLimit := 0.0;
   Machine[1].PneumaticFlow.PV_ActV.Value := 0.0;
   Machine[1].PneumaticFlow.PV_ActV.ValueState := 16#0000;
   Machine[1].PneumaticFlow.PV_Conf_ActV.OffsetSignal := 0;
   Machine[1].PneumaticFlow.PV_Conf_ActV.MaxSignalResolution := 0.0;
   Machine[2].PneumaticFlow.PV_SetV.Value := 0.0;
   Machine[2].PneumaticFlow.PV_SetV.WarningLowerLimit := 0.0;